// TIA Portal project "DATN" (V16) (continued)
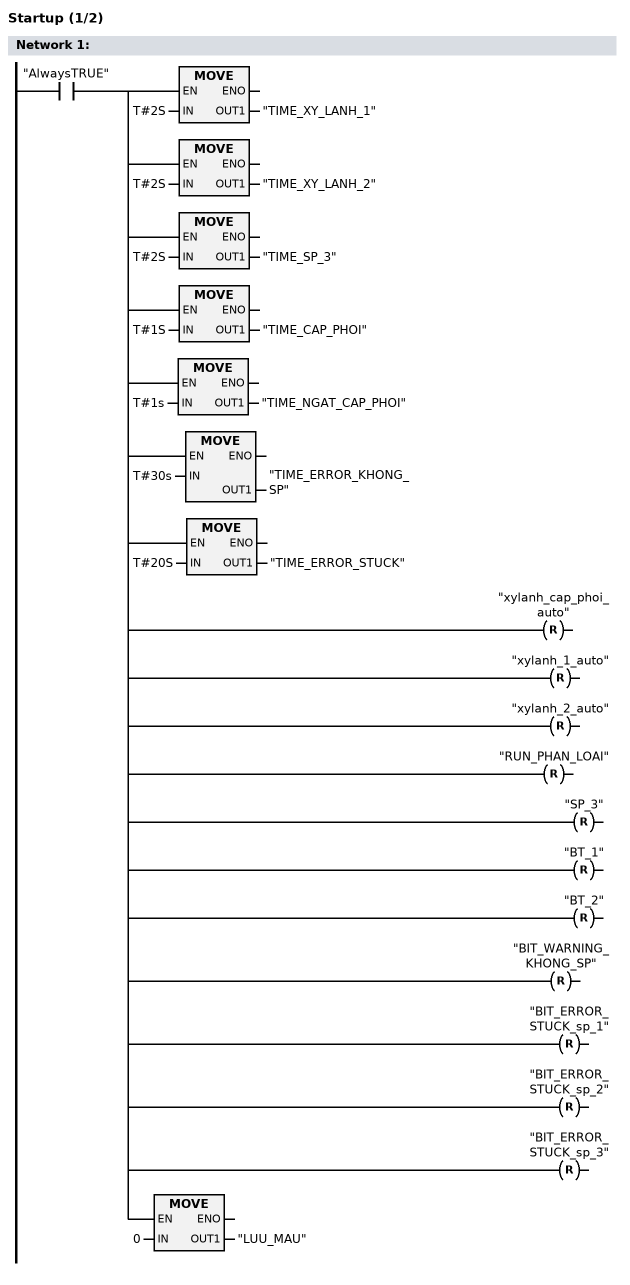
   RUNG wire#powerrail
      Contact( "AlwaysTRUE" )
      wire#w1
      Move(in := T#2S, out1 => "TIME_XY_LANH_1")
   END_RUNG
   RUNG wire#w1
      Move(in := T#2S, out1 => "TIME_XY_LANH_2")
   END_RUNG
   RUNG wire#w1
      Move(in := T#2S, out1 => "TIME_SP_3")
   END_RUNG
   RUNG wire#w1
      Move(in := T#1S, out1 => "TIME_CAP_PHOI")
   END_RUNG
   RUNG wire#w1
      Move(in := T#1s, out1 => "TIME_NGAT_CAP_PHOI")
   END_RUNG
   RUNG wire#w1
      Move(in := T#30s, out1 => "TIME_ERROR_KHONG_SP")
   END_RUNG
   RUNG wire#w1
      Move(in := T#20S, out1 => "TIME_ERROR_STUCK")
   END_RUNG
   RUNG wire#w1
      R_Coil( "xylanh_cap_phoi_auto" )
   END_RUNG
   RUNG wire#w1
      R_Coil( "xylanh_1_auto" )
   END_RUNG
   RUNG wire#w1
      R_Coil( "xylanh_2_auto" )
   END_RUNG
   RUNG wire#w1
      R_Coil( "RUN_PHAN_LOAI" )
   END_RUNG
   RUNG wire#w1
      R_Coil( "SP_3" )
   END_RUNG
   RUNG wire#w1
      R_Coil( "BT_1" )
   END_RUNG
   RUNG wire#w1
      R_Coil( "BT_2" )
   END_RUNG
   RUNG wire#w1
      R_Coil( "BIT_WARNING_KHONG_SP" )
   END_RUNG
   RUNG wire#w1
      R_Coil( "BIT_ERROR_STUCK_sp_1" )
   END_RUNG
   RUNG wire#w1
      R_Coil( "BIT_ERROR_STUCK_sp_2" )
   END_RUNG
   RUNG wire#w1
      R_Coil( "BIT_ERROR_STUCK_sp_3" )
   END_RUNG
   RUNG wire#w1
      Move(in := 0, out1 => "LUU_MAU")
   END_RUNG
   // the same network as SCL:
   IF "AlwaysTRUE" THEN
       "TIME_XY_LANH_1" := T#2S;
       "TIME_XY_LANH_2" := T#2S;
       "TIME_SP_3" := T#2S;
       "TIME_CAP_PHOI" := T#1S;
       "TIME_NGAT_CAP_PHOI" := T#1s;
       "TIME_ERROR_KHONG_SP" := T#30s;
       "TIME_ERROR_STUCK" := T#20S;
       "xylanh_cap_phoi_auto" := FALSE;
       "xylanh_1_auto" := FALSE;
       "xylanh_2_auto" := FALSE;
       "RUN_PHAN_LOAI" := FALSE;
       "SP_3" := FALSE;
       "BT_1" := FALSE;
       "BT_2" := FALSE;
       "BIT_WARNING_KHONG_SP" := FALSE;
       "BIT_ERROR_STUCK_sp_1" := FALSE;
       "BIT_ERROR_STUCK_sp_2" := FALSE;
       "BIT_ERROR_STUCK_sp_3" := FALSE;
       "LUU_MAU" := 0;
   END_IF;
END_REGION

REGION Network 2
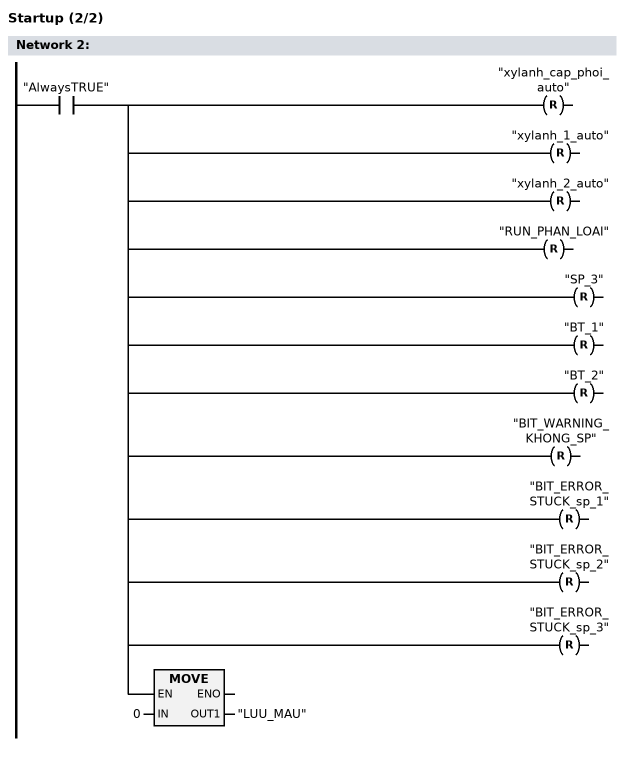
   RUNG wire#powerrail
      Contact( "AlwaysTRUE" )
      wire#w1
      R_Coil( "xylanh_cap_phoi_auto" )
   END_RUNG
   RUNG wire#w1
      R_Coil( "xylanh_1_auto" )
   END_RUNG
   RUNG wire#w1
      R_Coil( "xylanh_2_auto" )
   END_RUNG
   RUNG wire#w1
      R_Coil( "RUN_PHAN_LOAI" )
   END_RUNG
   RUNG wire#w1
      R_Coil( "SP_3" )
   END_RUNG
   RUNG wire#w1
      R_Coil( "BT_1" )
   END_RUNG
   RUNG wire#w1
      R_Coil( "BT_2" )
   END_RUNG
   RUNG wire#w1
      R_Coil( "BIT_WARNING_KHONG_SP" )
   END_RUNG
   RUNG wire#w1
      R_Coil( "BIT_ERROR_STUCK_sp_1" )
   END_RUNG
   RUNG wire#w1
      R_Coil( "BIT_ERROR_STUCK_sp_2" )
   END_RUNG
   RUNG wire#w1
      R_Coil( "BIT_ERROR_STUCK_sp_3" )
   END_RUNG
   RUNG wire#w1
      Move(in := 0, out1 => "LUU_MAU")
   END_RUNG
   // the same network as SCL:
   IF "AlwaysTRUE" THEN
       "xylanh_cap_phoi_auto" := FALSE;
       "xylanh_1_auto" := FALSE;
       "xylanh_2_auto" := FALSE;
       "RUN_PHAN_LOAI" := FALSE;
       "SP_3" := FALSE;
       "BT_1" := FALSE;
       "BT_2" := FALSE;
       "BIT_WARNING_KHONG_SP" := FALSE;
       "BIT_ERROR_STUCK_sp_1" := FALSE;
       "BIT_ERROR_STUCK_sp_2" := FALSE;
       "BIT_ERROR_STUCK_sp_3" := FALSE;
       "LUU_MAU" := 0;
   END_IF;
END_REGION
END_ORGANIZATION_BLOCK

(* ===== HMI "HMI_RT_1" =====
system functions are stored by id; their names below are inferred from use
connection "HMI_Connection_1": ETHERNET, S7_1200_OMS

HMI tags "Default tag table"
   "HMI_PB_START" : Bool = PLC HMI_PB_START AT %M100.4, 1 s
   "HMI_PB_STOP" : Bool = PLC HMI_PB_STOP AT %M100.5, 1 s
   "HMI_PB_RESET" : Bool = PLC HMI_PB_RESET AT %M100.6, 1 s
   "DEN_START" : Bool = PLC DEN_START AT %Q0.5, 1 s
   "DEN_STOP" : Bool = PLC DEN_STOP AT %Q0.6, 1 s
   "DEN_RESET" : Bool = PLC DEN_RESET AT %Q0.7, 1 s
   "HMI_AUTO_MAN" : Bool = PLC HMI_AUTO_MAN AT %M101.3, 1 s
   "COUNTER_SP_1_CV" : Int = PLC COUNTER_SP_1.CV, 1 s
   "COUNTER_SP_2_CV" : Int = PLC COUNTER_SP_2.CV, 1 s
   "COUNTER_SP_3_CV" : Int = PLC COUNTER_SP_3.CV, 1 s
   "gh_sp_GH_SP_1" : USInt = PLC gh_sp.GH_SP_1, 1 s
   "gh_sp_GH_SP_2" : USInt = PLC gh_sp.GH_SP_2, 1 s
   "gh_sp_GH_SP_3" : USInt = PLC gh_sp.GH_SP_3, 1 s
   "BANG_TAI" : Bool = PLC BANG_TAI AT %Q0.0, 1 s
   "XY_LANH_2" : Bool = PLC XY_LANH_2 AT %Q0.2, 1 s
   "XY_LANH_1" : Bool = PLC XY_LANH_1 AT %Q0.1, 1 s
   "Mau Sac" : Int = PLC "Mau Sac" AT %MW220, 1 s
   "CB_SP_2" : Bool = PLC CB_SP_2 AT %I0.2, 1 s
   "CB_SP_1" : Bool = PLC CB_SP_1 AT %I0.1, 1 s
   "CB_SP_3" : Bool = PLC CB_SP_3 AT %I0.3, 1 s
   "CB_CAP_PHOI" : Bool = PLC CB_CAP_PHOI AT %I0.0, 1 s
   "XY_LANH_CAP_PHOI_1" : Bool = PLC XY_LANH_CAP_PHOI_1 AT %Q0.3, 1 s
   "MODE_AUTO" : Bool = PLC MODE_AUTO AT %M201.7, 1 s
   "MODE_MAN" : Bool = PLC MODE_MAN AT %M202.0, 1 s
   "MAN_BT" : Bool = PLC MAN_BT AT %M100.7, 1 s
   "MAN_CAP_PHOI" : Bool = PLC MAN_CAP_PHOI AT %M101.2, 1 s
   "MAN_XYLANH_1" : Bool = PLC MAN_XYLANH_1 AT %M101.0, 1 s
   "MAN_XYLANH_2" : Bool = PLC MAN_XYLANH_2 AT %M101.1, 1 s
   "OUT_counter_1" : Bool = PLC OUT_counter_1 AT %M201.4, 1 s
   "OUT_counter_2" : Bool = PLC OUT_counter_2 AT %M201.5, 1 s
   "OUT_counter_3" : Bool = PLC OUT_counter_3 AT %M201.6, 1 s
   "RST_SP_3" : Bool = PLC RST_SP_3 AT %M101.6, 1 s
   "RST_SP_2" : Bool = PLC RST_SP_2 AT %M101.5, 1 s
   "RST_SP_1" : Bool = PLC RST_SP_1 AT %M101.4, 1 s
   "LUU_MAU" : Int = PLC LUU_MAU AT %MW222, 1 s
   "MULTI_ERROR" : Bool = PLC MULTI_ERROR AT %M450.0, 1 s
   "BIT_WARNING_KHONG_SP" : Bool = PLC BIT_WARNING_KHONG_SP AT %M400.0, 1 s
   "BIT_ERROR_STUCK_sp_1" : Bool = PLC BIT_ERROR_STUCK_sp_1 AT %M402.0, 1 s
   "BIT_ERROR_STUCK_sp_2" : Bool = PLC BIT_ERROR_STUCK_sp_2 AT %M404.0, 1 s
   "BIT_ERROR_STUCK_sp_3" : Bool = PLC BIT_ERROR_STUCK_sp_3 AT %M406.0, 1 s

HMI tags "HMI_ALARM"
   "DATA_WARNING" : Int = PLC DATA_WORD_WARNING AT %MW400, 1 s
   "DATA_ERROR_1" : Int = PLC DATA_WORD_ERROR_1 AT %MW402, 1 s
   "DATA_ERROR_2" : Int = PLC DATA_WORD_ERROR_2 AT %MW404, 1 s
   "DATA_ERROR_3" : Int = PLC DATA_WORD_ERROR_3 AT %MW406, 1 s

discrete alarms
   4: 'Cảnh báo không có sản phẩm', class Warnings, trigger "DATA_WARNING" bit 8
   1: 'Lỗi kẹt sản phẩm 1', class Warnings, trigger "DATA_ERROR_1" bit 8
   2: 'Lỗi kẹt sản phẩm 2', class Warnings, trigger "DATA_ERROR_2" bit 8
   3: 'Lỗi kẹt sản phẩm 3', class Warnings, trigger "DATA_ERROR_3" bit 8

screen "1_Login" 1440x900
   GraphicView "Graphic view_4" at 0,0 size 1438x897; Picture "plc"
   Button "Button_1" at 1010,602 size 237x78; TextOff 'LOG IN'; TextOn '2_Home'; Authorization "Operate"
      on Click: ActivateScreen("2_Home", 0)

screen "2_Home" 1440x900
   Circle "Circle_8" at 525,299 size 20x20
      Visibility <- "XY_LANH_2"
   Group "Group_7" at 531,249 size 89x62
   Polyline "Polyline_1" at 532,284 size 40x22
      Visibility <- "XY_LANH_2"
   Polyline "Polyline_2" at 531,249 size 89x62
      Visibility <- "XY_LANH_2"
   Group "Group_8" at 525,249 size 95x70
   Circle "Circle_9" at 525,299 size 20x20
      Visibility <- "XY_LANH_2"
   Circle "Circle_10" at 773,299 size 20x20
      Visibility <- "XY_LANH_1"
   Group "Group_9" at 779,249 size 89x62
   Polyline "Polyline_3" at 780,284 size 40x22
      Visibility <- "XY_LANH_1"
   Polyline "Polyline_4" at 779,249 size 89x62
      Visibility <- "XY_LANH_1"
   Group "Group_10" at 773,249 size 95x70
   Circle "Circle_11" at 773,299 size 20x20
      Visibility <- "XY_LANH_1"
   SymbolLibrary "Symbol library_14" at 1038,320 size 72x64
      Visibility <- "LUU_MAU"
   GraphicView "Graphic view_1" at 1039,340 size 58x29; Picture "Graphic_2"
      Visibility <- "LUU_MAU"
   SymbolLibrary "Symbol library_13" at 1020,330 size 72x64
      Visibility <- "LUU_MAU"
   GraphicView "Graphic view_3" at 1021,348 size 58x33; Picture "Graphic_4"
      Visibility <- "LUU_MAU"
   SymbolLibrary "Symbol library_12" at 1002,342 size 72x64
      Visibility <- "LUU_MAU"
   GraphicView "Graphic view_2" at 1003,360 size 58x33; Picture "Graphic_5"
      Visibility <- "LUU_MAU"
   SymbolLibrary "Symbol library_21" at 349,368 size 17x150
   SymbolLibrary "Symbol library_6" at 93,426 size 168x95
      Appearance <- "OUT_counter_3"
   SymbolLibrary "Symbol library_17" at 333,345 size 56x52
   SymbolLibrary "Symbol library_20" at 1179,373 size 17x150
   SymbolLibrary "Symbol library_16" at 1161,350 size 56x52
   SymbolLibrary "Symbol library_1" at 242,368 size 545x73
      Appearance <- "BANG_TAI"
   SymbolLibrary "Symbol library_2" at 650,368 size 545x73
      Appearance <- "BANG_TAI"
   SymbolLibrary "Symbol library_19" at 1082,432 size 17x150
   Group "Group_6" at 595,168 size 143x104
   Group "Group_12" at 525,249 size 95x70
   Group "Group_1" at 843,168 size 143x104
   Group "Group_11" at 773,249 size 95x70
   SymbolLibrary "Symbol library_4" at 334,546 size 168x95
      Appearance <- "OUT_counter_2"
   SymbolLibrary "Symbol library_5" at 570,546 size 168x95
      Appearance <- "OUT_counter_1"
   SymbolLibrary "Symbol library_8" at 1025,248 size 55x27
      Appearance <- "Mau Sac"
   SymbolLibrary "Symbol library_10" at 649,242 size 28x55
      Appearance <- "CB_SP_2"
   SymbolLibrary "Symbol library_11" at 902,242 size 28x55
      Appearance <- "CB_SP_1"
   TextField "Text field_6" at 679,244 size 39x25; Text 'CB2'
   TextField "Text field_7" at 931,244 size 39x25; Text 'CB1'
   TextField "Text field_9" at 569,140 size 114x56; Text 'Xy lanh loại 2'
   TextField "Text field_10" at 826,140 size 114x56; Text 'Xy lanh loại 1'
   IOField "I/O field_4" at 378,594 size 62x32; FormatPattern 99999
      ProcessValue <- "COUNTER_SP_2_CV"
   IOField "I/O field_5" at 614,594 size 62x32; FormatPattern 99999
      ProcessValue <- "COUNTER_SP_1_CV"
   TextField "Text field_14" at 103,514 size 123x43; Text 'SP Loại 3'
   TextField "Text field_15" at 456,605 size 123x43; Text 'SP Loại 2'
   TextField "Text field_16" at 693,605 size 123x43; Text 'SP Loại 1'
   Group "Group_15" at 1038,320 size 72x64; Picture "Graphic_2"
   Group "Group_16" at 1020,330 size 72x64; Picture "Graphic_4"
   SymbolLibrary "Symbol library_15" at 1065,403 size 56x52
   TextField "Text field_17" at 899,520 size 138x61; Text 'ĐỘNG CƠ BĂNG TẢI'
   Group "Group_17" at 1002,342 size 72x64; Picture "Graphic_5"
   Group "Group_13" at 385,415 size 133x122
   SymbolLibrary "Symbol library_3" at 928,463 size 110x66
      Appearance <- "BANG_TAI"
   IOField "I/O field_6" at 137,480 size 62x32; FormatPattern 99999
      ProcessValue <- "COUNTER_SP_3_CV"
   SymbolLibrary "Symbol library_22" at 243,427 size 17x150
   SymbolLibrary "Symbol library_18" at 225,404 size 56x52
   Group "Group_2" at 625,415 size 133x122
   Button "Button_3" at 11,123 size 112x37; TextOff 'Home'
      on Click: ActivateScreen("2_Home", 0)
   Button "Button_4" at 11,177 size 112x37; TextOff 'Control'; Authorization "User administration"
      on Click: ActivateScreen("3_Control", 0)
   Button "Button_6" at 11,285 size 112x37; TextOff 'Log out'
      on Click: function_f23ef4c9(); ActivateScreen("1_Login", 0)
   DateTimeField "Date/time field_3" at 1186,44 size 102x23
   DateTimeField "Date/time field_1" at 1186,18 size 254x23
   GraphicView "Graphic view_8" at 38,8 size 70x70; Picture "Hcmute"
   GraphicView "Graphic view_9" at 128,8 size 70x70; Picture "feee"
   TextField "Text field_3" at 261,15 size 906x70; Text 'HỆ THỐNG PHÂN LOẠI SẢN PHẨM THEO MÀU SẮC DÙNG XỬ LÝ ẢNH'
   GraphicView "Graphic view_10" at 134,130 size 36x18; Picture "Graphic_17"
   TextField "Text field_1" at 250,147 size 15x22; Text 'Text'
   TextField "Text field_4" at 72,730 size 139x22; Text 'Hệ thống nút nhấn'
   Button "Button_1" at 26,801 size 64x64; TextOff 'Text'; PictureOff "3-D green button (not pressed)_3"; PictureOn "3-D green button (pressed)_2"
      on Press: SetBit("HMI_PB_START")
      on Release: ResetBit("HMI_PB_START")
   TextField "Text field_5" at 31,768 size 54x22; Text 'START'
   TextField "Text field_8" at 353,730 size 133x22; Text 'Hệ thống đèn báo'
   Button "Button_2" at 109,801 size 64x64; TextOff 'Text'; PictureOff "3-D red button (not pressed)"; PictureOn "3-D red button (pressed)"
      on Press: SetBit("HMI_PB_STOP")
      on Release: ResetBit("HMI_PB_STOP")
   TextField "Text field_11" at 118,768 size 46x22; Text 'STOP'
   Button "Button_7" at 193,801 size 64x64; TextOff 'Text'; PictureOff "3-D yellow button (not pressed)"; PictureOn "3-D yellow button (pressed)"
      on Press: SetBit("HMI_PB_RESET")
      on Release: ResetBit("HMI_PB_RESET")
   TextField "Text field_12" at 199,768 size 53x22; Text 'RESET'
   GraphicView "Graphic view_4" at 387,801 size 64x64; Picture "Graphic_11"
      Visibility <- "DEN_STOP"
   GraphicView "Graphic view_5" at 304,801 size 64x64; Picture "Graphic_9"
      Visibility <- "DEN_START"
   GraphicView "Graphic view_6" at 471,801 size 64x64; Picture "Graphic_18"
      Visibility <- "DEN_RESET"
   GraphicView "Graphic view_7" at 304,801 size 64x64; Picture "Graphic_10"
      Visibility <- "DEN_START"
   GraphicView "Graphic view_11" at 387,801 size 64x64; Picture "Graphic_12"
      Visibility <- "DEN_STOP"
   GraphicView "Graphic view_12" at 471,801 size 64x64; Picture "Graphic_19"
      Visibility <- "DEN_RESET"
   TextField "Text field_13" at 322,768 size 29x22; Text 'ON'
   TextField "Text field_18" at 402,768 size 35x22; Text 'OFF'
   TextField "Text field_19" at 456,768 size 95x22; Text 'WARNNING'
   TextField "Text field_20" at 659,683 size 123x22; Text 'Bảng điều khiển'
   TextField "Text field_2" at 581,730 size 132x22; Text 'Chế độ hoạt động'
   Switch "Switch_1" at 587,805 size 120x60; CaptionText 'Switch'; TextOff 'OFF'; TextOn 'ON'; PictureOn "Illuminated red-green (Red)_1"; PictureOff "Illuminated red-green (Green)_1"
      ProcessValue <- "HMI_AUTO_MAN"
   TextField "Text field_23" at 973,730 size 148x22; Text 'Thông tin sản phẩm'
   TextField "Text field_24" at 895,754 size 137x22; Text 'Giới hạn số lượng'
   TextField "Text field_25" at 760,784 size 123x22; Text 'Sản phẩm loại 1'
   TextField "Text field_26" at 760,816 size 123x22; Text 'Sản phẩm loại 2'
   TextField "Text field_27" at 760,848 size 123x22; Text 'Sản phẩm loại 3'
   IOField "I/O field_1" at 916,779 size 96x32; FormatPattern 999
      ProcessValue <- "gh_sp_GH_SP_1"
   IOField "I/O field_2" at 916,811 size 96x32; FormatPattern 999
      ProcessValue <- "gh_sp_GH_SP_2"
   IOField "I/O field_3" at 916,843 size 96x32; FormatPattern 999
      ProcessValue <- "gh_sp_GH_SP_3"
   TextField "Text field_28" at 1084,754 size 130x22; Text 'Số lượng hiện tại'
   IOField "I/O field_7" at 1101,779 size 96x32; FormatPattern 99999
      ProcessValue <- "COUNTER_SP_1_CV"
   IOField "I/O field_8" at 1101,811 size 96x32; FormatPattern 99999
      ProcessValue <- "COUNTER_SP_2_CV"
   IOField "I/O field_9" at 1101,843 size 96x32; FormatPattern 99999
      ProcessValue <- "COUNTER_SP_3_CV"
   GraphicView "Graphic view_13" at 1023,406 size 94x98; Picture "Graphic_20"
   SymbolLibrary "Symbol library_7" at 349,242 size 28x55
      Appearance <- "CB_SP_3"
   TextField "Text field_29" at 385,244 size 39x25; Text 'CB3'
   SymbolLibrary "Symbol library_23" at 1215,367 size 17x155
   SymbolLibrary "Symbol library_24" at 1118,426 size 17x156
   SymbolLibrary "Symbol library_25" at 1302,367 size 17x154
   SymbolLibrary "Symbol library_26" at 1205,426 size 17x155
   SymbolLibrary "Symbol library_27" at 1183,330 size 72x64
      Visibility <- "CB_CAP_PHOI"
   SymbolLibrary "Symbol library_28" at 1287,316 size 55x28
      Appearance <- "CB_CAP_PHOI"
   SymbolLibrary "Symbol library_9" at 1243,351 size 130x26
      Visibility <- "XY_LANH_CAP_PHOI_1"
   SymbolLibrary "Symbol library_29" at 1292,351 size 82x26
      Visibility <- "XY_LANH_CAP_PHOI_1"
   TextField "Text field_30" at 1270,281 size 117x25; Text 'CB CẤP PHÔI'
   TextField "Text field_31" at 1258,754 size 134x22; Text 'Reset thùng hàng'
   Button "Button_8" at 1277,779 size 96x32; TextOff 'RST_1'
      Appearance <- "OUT_counter_1"
      on Press: SetBit("RST_SP_1")
      on Release: ResetBit("RST_SP_1")
   Button "Button_9" at 1277,810 size 96x32; TextOff 'RST_2'
      Appearance <- "OUT_counter_2"
      on Press: SetBit("RST_SP_2")
      on Release: ResetBit("RST_SP_2")
   Button "Button_10" at 1277,841 size 96x32; TextOff 'RST_3'
      Appearance <- "OUT_counter_3"
      on Press: SetBit("RST_SP_3")
      on Release: ResetBit("RST_SP_3")
   Button "Button_5" at 11,231 size 112x37; TextOff 'Alarm'
      on Click: ActivateScreen("4_ALARM", 0)
      Appearance <- "MULTI_ERROR"
   Rectangle "Rectangle_9" at 579,754 size 65x48
      Appearance <- "MODE_AUTO"
   Rectangle "Rectangle_10" at 650,754 size 65x48
      Appearance <- "MODE_MAN"
   TextField "Text field_32" at 1203,96 size 125x22; Text 'Màu sắc hiện tại'
   Rectangle "Rectangle_13" at 1246,137 size 40x37
      Appearance <- "LUU_MAU"
   TextField "Text field_33" at 1245,185 size 42x22; Text 'Vàng'
      Visibility <- "LUU_MAU"
   TextField "Text field_34" at 1248,185 size 36x22; Text 'Lam'
      Visibility <- "LUU_MAU"
   TextField "Text field_35" at 1250,185 size 32x22; Text 'Tím'
      Visibility <- "LUU_MAU"
   TextField "Text field_36" at 1231,185 size 70x22; Text 'No Color'
      Visibility <- "LUU_MAU"
   TextField "Text field_21" at 592,768 size 39x22; Text 'Auto'
   TextField "Text field_22" at 653,768 size 59x22; Text 'Manual'

screen "3_Control" 1440x900
   Circle "Circle_8" at 525,299 size 20x20
      Visibility <- "XY_LANH_2"
   Group "Group_7" at 531,249 size 89x62
   Polyline "Polyline_1" at 532,284 size 40x22
      Visibility <- "XY_LANH_2"
   Polyline "Polyline_2" at 531,249 size 89x62
      Visibility <- "XY_LANH_2"
   Group "Group_8" at 525,249 size 95x70
   Circle "Circle_9" at 525,299 size 20x20
      Visibility <- "XY_LANH_2"
   Circle "Circle_10" at 773,299 size 20x20
      Visibility <- "XY_LANH_1"
   Group "Group_9" at 779,249 size 89x62
   Polyline "Polyline_3" at 780,284 size 40x22
      Visibility <- "XY_LANH_1"
   Polyline "Polyline_4" at 779,249 size 89x62
      Visibility <- "XY_LANH_1"
   Group "Group_10" at 773,249 size 95x70
   Circle "Circle_11" at 773,299 size 20x20
      Visibility <- "XY_LANH_1"
   SymbolLibrary "Symbol library_6" at 93,426 size 168x95
      Appearance <- "OUT_counter_3"
   SymbolLibrary "Symbol library_4" at 334,546 size 168x95
      Appearance <- "OUT_counter_2"
   SymbolLibrary "Symbol library_5" at 570,546 size 168x95
      Appearance <- "OUT_counter_1"
   SymbolLibrary "Symbol library_21" at 349,368 size 17x150
   SymbolLibrary "Symbol library_17" at 333,345 size 56x52
   SymbolLibrary "Symbol library_20" at 1179,373 size 17x150
   SymbolLibrary "Symbol library_16" at 1161,350 size 56x52
   SymbolLibrary "Symbol library_1" at 242,368 size 545x73
      Appearance <- "BANG_TAI"
   SymbolLibrary "Symbol library_2" at 650,368 size 545x73
      Appearance <- "BANG_TAI"
   SymbolLibrary "Symbol library_19" at 1082,432 size 17x150
   Group "Group_6" at 595,168 size 143x104
   Group "Group_12" at 525,249 size 95x70
   Group "Group_1" at 843,168 size 143x104
   Group "Group_11" at 773,249 size 95x70
   SymbolLibrary "Symbol library_8" at 1025,248 size 55x27
      Appearance <- "Mau Sac"
   SymbolLibrary "Symbol library_10" at 649,242 size 28x55
      Appearance <- "CB_SP_2"
   SymbolLibrary "Symbol library_11" at 902,242 size 28x55
      Appearance <- "CB_SP_1"
   TextField "Text field_6" at 679,244 size 39x25; Text 'CB2'
   TextField "Text field_7" at 931,244 size 39x25; Text 'CB1'
   TextField "Text field_9" at 569,140 size 114x56; Text 'Xy lanh loại 2'
   TextField "Text field_10" at 826,140 size 114x56; Text 'Xy lanh loại 1'
   IOField "I/O field_4" at 378,594 size 62x32; FormatPattern 99999
      ProcessValue <- "COUNTER_SP_2_CV"
   IOField "I/O field_5" at 614,594 size 62x32; FormatPattern 99999
      ProcessValue <- "COUNTER_SP_1_CV"
   TextField "Text field_14" at 103,514 size 123x43; Text 'SP Loại 3'
   TextField "Text field_15" at 456,605 size 123x43; Text 'SP Loại 2'
   TextField "Text field_16" at 693,605 size 123x43; Text 'SP Loại 1'
   SymbolLibrary "Symbol library_15" at 1065,403 size 56x52
   TextField "Text field_17" at 899,520 size 138x61; Text 'ĐỘNG CƠ BĂNG TẢI'
   Group "Group_13" at 385,415 size 133x122
   SymbolLibrary "Symbol library_3" at 928,463 size 110x66
      Appearance <- "BANG_TAI"
   IOField "I/O field_6" at 137,480 size 62x32; FormatPattern 99999
      ProcessValue <- "COUNTER_SP_3_CV"
   SymbolLibrary "Symbol library_22" at 243,427 size 17x150
   SymbolLibrary "Symbol library_18" at 225,404 size 56x52
   Group "Group_2" at 625,415 size 133x122
   Button "Button_3" at 11,123 size 112x37; TextOff 'Home'
      on Click: ActivateScreen("2_Home", 0)
   Button "Button_4" at 11,177 size 112x37; TextOff 'Control'
      on Click: ActivateScreen("3_Control", 0)
   Button "Button_6" at 11,285 size 112x37; TextOff 'Log out'
      on Click: ActivateScreen("1_Login", 0)
   DateTimeField "Date/time field_3" at 1186,44 size 102x23
   DateTimeField "Date/time field_1" at 1186,18 size 254x23
   GraphicView "Graphic view_8" at 38,8 size 70x70; Picture "Hcmute"
   GraphicView "Graphic view_9" at 128,8 size 70x70; Picture "feee"
   GraphicView "Graphic view_10" at 134,187 size 36x18; Picture "Graphic_17"
   TextField "Text field_1" at 250,147 size 15x22; Text 'Text'
   TextField "Text field_4" at 72,730 size 139x22; Text 'Hệ thống nút nhấn'
   Button "Button_1" at 26,801 size 64x64; TextOff 'Text'; PictureOn "3-D green button (pressed)_2"; PictureOff "3-D green button (not pressed)_3"
      on Release: ResetBit("HMI_PB_START")
      on Press: SetBit("HMI_PB_START")
   TextField "Text field_5" at 31,768 size 54x22; Text 'START'
   TextField "Text field_8" at 353,730 size 133x22; Text 'Hệ thống đèn báo'
   Button "Button_2" at 109,801 size 64x64; TextOff 'Text'; PictureOn "3-D red button (pressed)"; PictureOff "3-D red button (not pressed)"
      on Release: ResetBit("HMI_PB_STOP")
      on Press: SetBit("HMI_PB_STOP")
   TextField "Text field_11" at 118,768 size 46x22; Text 'STOP'
   Button "Button_7" at 193,801 size 64x64; TextOff 'Text'; PictureOn "3-D yellow button (pressed)"; PictureOff "3-D yellow button (not pressed)"
      on Release: ResetBit("HMI_PB_RESET")
      on Press: SetBit("HMI_PB_RESET")
   TextField "Text field_12" at 199,768 size 53x22; Text 'RESET'
   GraphicView "Graphic view_4" at 387,801 size 64x64; Picture "Graphic_11"
      Visibility <- "DEN_STOP"
   GraphicView "Graphic view_5" at 304,801 size 64x64; Picture "Graphic_9"
      Visibility <- "DEN_START"
   GraphicView "Graphic view_6" at 471,801 size 64x64; Picture "Graphic_18"
      Visibility <- "DEN_RESET"
   GraphicView "Graphic view_7" at 304,801 size 64x64; Picture "Graphic_10"
      Visibility <- "DEN_START"
   GraphicView "Graphic view_11" at 387,801 size 64x64; Picture "Graphic_12"
      Visibility <- "DEN_STOP"
   GraphicView "Graphic view_12" at 471,801 size 64x64; Picture "Graphic_19"
      Visibility <- "DEN_RESET"
   TextField "Text field_13" at 322,768 size 29x22; Text 'ON'
   TextField "Text field_18" at 402,768 size 35x22; Text 'OFF'
   TextField "Text field_19" at 456,768 size 95x22; Text 'WARNNING'
   TextField "Text field_20" at 659,683 size 123x22; Text 'Bảng điều khiển'
   TextField "Text field_2" at 581,730 size 132x22; Text 'Chế độ hoạt động'
   Switch "Switch_1" at 587,805 size 120x60; CaptionText 'Switch'; TextOff 'OFF'; TextOn 'ON'; PictureOff "Illuminated red-green (Green)_1"; PictureOn "Illuminated red-green (Red)_1"
      ProcessValue <- "HMI_AUTO_MAN"
   TextField "Text field_23" at 746,730 size 261x22; Text 'Cài đặt giới hạn số lượng sản phẩm'
   TextField "Text field_25" at 745,784 size 123x22; Text 'Sản phẩm loại 1'
   TextField "Text field_26" at 745,816 size 123x22; Text 'Sản phẩm loại 2'
   TextField "Text field_27" at 745,848 size 123x22; Text 'Sản phẩm loại 3'
   IOField "I/O field_1" at 901,779 size 96x32; FormatPattern 999
      ProcessValue <- "gh_sp_GH_SP_1"
   IOField "I/O field_2" at 901,811 size 96x32; FormatPattern 999
      ProcessValue <- "gh_sp_GH_SP_2"
   IOField "I/O field_3" at 901,843 size 96x32; FormatPattern 999
      ProcessValue <- "gh_sp_GH_SP_3"
   GraphicView "Graphic view_13" at 1023,406 size 94x98; Picture "Graphic_20"
   SymbolLibrary "Symbol library_7" at 349,242 size 28x55
      Appearance <- "CB_SP_3"
   TextField "Text field_29" at 385,244 size 39x25; Text 'CB3'
   SymbolLibrary "Symbol library_23" at 1215,367 size 17x155
   SymbolLibrary "Symbol library_24" at 1118,426 size 17x156
   SymbolLibrary "Symbol library_25" at 1302,367 size 17x154
   SymbolLibrary "Symbol library_26" at 1205,426 size 17x155
   SymbolLibrary "Symbol library_27" at 1183,330 size 72x64
      Visibility <- "CB_CAP_PHOI"
   SymbolLibrary "Symbol library_28" at 1287,316 size 55x28
      Appearance <- "CB_CAP_PHOI"
   SymbolLibrary "Symbol library_9" at 1243,351 size 130x26
      Visibility <- "XY_LANH_CAP_PHOI_1"
   SymbolLibrary "Symbol library_29" at 1292,351 size 82x26
      Visibility <- "XY_LANH_CAP_PHOI_1"
   TextField "Text field_30" at 1270,281 size 117x25; Text 'CB CẤP PHÔI'
   Rectangle "Rectangle_9" at 579,754 size 65x48
      Appearance <- "MODE_AUTO"
   Rectangle "Rectangle_10" at 650,754 size 65x48
      Appearance <- "MODE_MAN"
   TextField "Text field_21" at 592,768 size 39x22; Text 'Auto'
   TextField "Text field_22" at 653,768 size 59x22; Text 'Manual'
   TextField "Text field_24" at 1158,730 size 153x22; Text 'Điều khiển bằng tay'
   Button "Button_8" at 1062,779 size 160x32; TextOff 'Băng tải'
      Appearance <- "BANG_TAI"
      on Press: SetBit("MAN_BT")
      on Release: ResetBit("MAN_BT")
   Button "Button_9" at 1062,843 size 160x32; TextOff 'Xylanh cấp phôi'
      Appearance <- "XY_LANH_CAP_PHOI_1"
      on Press: SetBit("MAN_CAP_PHOI")
      on Release: ResetBit("MAN_CAP_PHOI")
   Button "Button_10" at 1256,779 size 160x32; TextOff 'Xylanh 1'
      Appearance <- "XY_LANH_1"
      on Press: SetBit("MAN_XYLANH_1")
      on Release: ResetBit("MAN_XYLANH_1")
   Button "Button_11" at 1256,843 size 160x32; TextOff 'Xylanh 2'
      Appearance <- "XY_LANH_2"
      on Press: SetBit("MAN_XYLANH_2")
      on Release: ResetBit("MAN_XYLANH_2")
   Button "Button_5" at 11,231 size 112x37; TextOff 'Alarm'
      on Click: ActivateScreen("4_ALARM", 0)
      Appearance <- "MULTI_ERROR"
   TextField "Text field_32" at 1203,96 size 125x22; Text 'Màu sắc hiện tại'
   Rectangle "Rectangle_13" at 1246,137 size 40x37
      Appearance <- "LUU_MAU"
   TextField "Text field_33" at 1245,185 size 42x22; Text 'Vàng'
      Visibility <- "LUU_MAU"
   TextField "Text field_34" at 1248,185 size 36x22; Text 'Lam'
      Visibility <- "LUU_MAU"
   TextField "Text field_35" at 1250,185 size 32x22; Text 'Tím'
      Visibility <- "LUU_MAU"
   TextField "Text field_36" at 1231,185 size 70x22; Text 'No Color'
      Visibility <- "LUU_MAU"
   Group "Group_15" at 1038,320 size 72x64; Picture "Graphic_2"
   Group "Group_16" at 1020,330 size 72x64; Picture "Graphic_4"
   Group "Group_17" at 1002,342 size 72x64; Picture "Graphic_5"
   TextField "Text field_3" at 261,15 size 906x70; Text 'HỆ THỐNG PHÂN LOẠI SẢN PHẨM THEO MÀU SẮC DÙNG XỬ LÝ ẢNH'
   SymbolLibrary "Symbol library_14" at 1038,320 size 72x64
      Visibility <- "LUU_MAU"
   GraphicView "Graphic view_1" at 1039,340 size 58x29; Picture "Graphic_2"
      Visibility <- "LUU_MAU"
   SymbolLibrary "Symbol library_13" at 1020,330 size 72x64
      Visibility <- "LUU_MAU"
   GraphicView "Graphic view_3" at 1021,348 size 58x33; Picture "Graphic_4"
      Visibility <- "LUU_MAU"
   SymbolLibrary "Symbol library_12" at 1002,342 size 72x64
      Visibility <- "LUU_MAU"
   GraphicView "Graphic view_2" at 1003,360 size 58x33; Picture "Graphic_5"
      Visibility <- "LUU_MAU"

screen "4_ALARM" 1440x900
   SymbolLibrary "Symbol library_21" at 349,368 size 17x150
   SymbolLibrary "Symbol library_6" at 93,426 size 168x95
      Appearance <- "OUT_counter_3"
   SymbolLibrary "Symbol library_17" at 333,345 size 56x52
   SymbolLibrary "Symbol library_20" at 1179,373 size 17x150
   SymbolLibrary "Symbol library_16" at 1161,350 size 56x52
   SymbolLibrary "Symbol library_1" at 242,368 size 545x73
      Appearance <- "BANG_TAI"
   SymbolLibrary "Symbol library_2" at 650,368 size 545x73
      Appearance <- "BANG_TAI"
   SymbolLibrary "Symbol library_19" at 1082,432 size 17x150
   Group "Group_6" at 595,168 size 143x104
   Group "Group_12" at 525,249 size 95x70
   Group "Group_1" at 843,168 size 143x104
   Group "Group_11" at 773,249 size 95x70
   SymbolLibrary "Symbol library_4" at 334,546 size 168x95
      Appearance <- "OUT_counter_2"
   SymbolLibrary "Symbol library_5" at 570,546 size 168x95
      Appearance <- "OUT_counter_1"
   SymbolLibrary "Symbol library_8" at 1025,248 size 55x27
      Appearance <- "Mau Sac"
   SymbolLibrary "Symbol library_10" at 649,242 size 28x55
      Appearance <- "CB_SP_2"
   SymbolLibrary "Symbol library_11" at 902,242 size 28x55
      Appearance <- "CB_SP_1"
   TextField "Text field_6" at 679,244 size 39x25; Text 'CB2'
   TextField "Text field_7" at 931,244 size 39x25; Text 'CB1'
   TextField "Text field_9" at 569,140 size 114x56; Text 'Xy lanh loại 2'
   TextField "Text field_10" at 826,140 size 114x56; Text 'Xy lanh loại 1'
   IOField "I/O field_4" at 378,594 size 62x32; FormatPattern 99999
      ProcessValue <- "COUNTER_SP_2_CV"
   IOField "I/O field_5" at 614,594 size 62x32; FormatPattern 99999
      ProcessValue <- "COUNTER_SP_1_CV"
   TextField "Text field_14" at 103,514 size 123x43; Text 'SP Loại 3'
   TextField "Text field_15" at 456,605 size 123x43; Text 'SP Loại 2'
   TextField "Text field_16" at 693,605 size 123x43; Text 'SP Loại 1'
   SymbolLibrary "Symbol library_15" at 1065,403 size 56x52
   TextField "Text field_17" at 899,520 size 138x61; Text 'ĐỘNG CƠ BĂNG TẢI'
   Group "Group_13" at 385,415 size 133x122
   SymbolLibrary "Symbol library_3" at 928,463 size 110x66
      Appearance <- "BANG_TAI"
   IOField "I/O field_6" at 137,480 size 62x32; FormatPattern 99999
      ProcessValue <- "COUNTER_SP_3_CV"
   SymbolLibrary "Symbol library_22" at 243,427 size 17x150
   SymbolLibrary "Symbol library_18" at 225,404 size 56x52
   Group "Group_2" at 625,415 size 133x122
   Button "Button_3" at 11,123 size 112x37; TextOff 'Home'
      on Click: ActivateScreen("2_Home", 0)
   Button "Button_4" at 11,177 size 112x37; TextOff 'Control'
      on Click: ActivateScreen("3_Control", 0)
   Button "Button_5" at 11,231 size 112x37; TextOff 'Alarm'
      on Click: ActivateScreen("4_ALARM", 0)
      Appearance <- "MULTI_ERROR"
   Button "Button_6" at 11,285 size 112x37; TextOff 'Log out'
      on Click: function_f23ef4c9(); ActivateScreen("1_Login", 0)
   DateTimeField "Date/time field_3" at 1186,44 size 102x23
   DateTimeField "Date/time field_1" at 1186,18 size 254x23
   GraphicView "Graphic view_8" at 38,8 size 70x70; Picture "Hcmute"
   GraphicView "Graphic view_9" at 128,8 size 70x70; Picture "feee"
   GraphicView "Graphic view_10" at 134,241 size 36x18; Picture "Graphic_17"
   TextField "Text field_1" at 250,147 size 15x22; Text 'Text'
   TextField "Text field_4" at 72,730 size 139x22; Text 'Hệ thống nút nhấn'
   Button "Button_1" at 26,801 size 64x64; TextOff 'Text'; PictureOn "3-D green button (pressed)_2"; PictureOff "3-D green button (not pressed)_3"
      on Release: ResetBit("HMI_PB_START")
      on Press: SetBit("HMI_PB_START")
   TextField "Text field_5" at 31,768 size 54x22; Text 'START'
   TextField "Text field_8" at 353,730 size 133x22; Text 'Hệ thống đèn báo'
   Button "Button_2" at 109,801 size 64x64; TextOff 'Text'; PictureOn "3-D red button (pressed)"; PictureOff "3-D red button (not pressed)"
      on Release: ResetBit("HMI_PB_STOP")
      on Press: SetBit("HMI_PB_STOP")
   TextField "Text field_11" at 118,768 size 46x22; Text 'STOP'
   Button "Button_7" at 193,801 size 64x64; TextOff 'Text'; PictureOn "3-D yellow button (pressed)"; PictureOff "3-D yellow button (not pressed)"
      on Release: ResetBit("HMI_PB_RESET")
      on Press: SetBit("HMI_PB_RESET")
   TextField "Text field_12" at 199,768 size 53x22; Text 'RESET'
   GraphicView "Graphic view_4" at 387,801 size 64x64; Picture "Graphic_11"
      Visibility <- "DEN_STOP"
   GraphicView "Graphic view_5" at 304,801 size 64x64; Picture "Graphic_9"
      Visibility <- "DEN_START"
   GraphicView "Graphic view_6" at 471,801 size 64x64; Picture "Graphic_18"
      Visibility <- "DEN_RESET"
   GraphicView "Graphic view_7" at 304,801 size 64x64; Picture "Graphic_10"
      Visibility <- "DEN_START"
   GraphicView "Graphic view_11" at 387,801 size 64x64; Picture "Graphic_12"
      Visibility <- "DEN_STOP"
   GraphicView "Graphic view_12" at 471,801 size 64x64; Picture "Graphic_19"
      Visibility <- "DEN_RESET"
   TextField "Text field_13" at 322,768 size 29x22; Text 'ON'
   TextField "Text field_18" at 402,768 size 35x22; Text 'OFF'
   TextField "Text field_19" at 456,768 size 95x22; Text 'WARNNING'
   TextField "Text field_20" at 659,683 size 123x22; Text 'Bảng điều khiển'
   TextField "Text field_2" at 581,730 size 132x22; Text 'Chế độ hoạt động'
   Switch "Switch_1" at 587,805 size 120x60; CaptionText 'Switch'; TextOff 'OFF'; TextOn 'ON'; PictureOff "Illuminated red-green (Green)_1"; PictureOn "Illuminated red-green (Red)_1"
      ProcessValue <- "HMI_AUTO_MAN"
   GraphicView "Graphic view_13" at 1023,406 size 94x98; Picture "Graphic_20"
   SymbolLibrary "Symbol library_7" at 349,242 size 28x55
      Appearance <- "CB_SP_3"
   TextField "Text field_29" at 385,244 size 39x25; Text 'CB3'
   SymbolLibrary "Symbol library_23" at 1215,367 size 17x155
   SymbolLibrary "Symbol library_24" at 1118,426 size 17x156
   SymbolLibrary "Symbol library_25" at 1302,367 size 17x154
   SymbolLibrary "Symbol library_26" at 1205,426 size 17x155
   Polygon "Polygon_5" at 1118,366 size 202x60
      Appearance <- "BIT_WARNING_KHONG_SP"
   SymbolLibrary "Symbol library_27" at 1183,330 size 72x64
      Visibility <- "CB_CAP_PHOI"
   SymbolLibrary "Symbol library_28" at 1287,316 size 55x28
      Appearance <- "CB_CAP_PHOI"
   SymbolLibrary "Symbol library_9" at 1243,351 size 130x26
      Visibility <- "XY_LANH_CAP_PHOI_1"
   SymbolLibrary "Symbol library_29" at 1292,351 size 82x26
      Visibility <- "XY_LANH_CAP_PHOI_1"
   TextField "Text field_30" at 1270,281 size 117x25; Text 'CB CẤP PHÔI'
   AlarmView "Alarm view_1" at 739,716 size 680x169
   Rectangle "Rectangle_9" at 579,754 size 65x48
      Appearance <- "MODE_AUTO"
   Rectangle "Rectangle_10" at 650,754 size 65x48
      Appearance <- "MODE_MAN"
   TextField "Text field_21" at 592,768 size 39x22; Text 'Auto'
   TextField "Text field_22" at 653,768 size 59x22; Text 'Manual'
   Group "Group_3" at 882,342 size 72x64; Picture "Graphic_5"
   TextField "Text field_32" at 1203,96 size 125x22; Text 'Màu sắc hiện tại'
   Rectangle "Rectangle_13" at 1246,137 size 40x37
      Appearance <- "LUU_MAU"
   TextField "Text field_33" at 1245,185 size 42x22; Text 'Vàng'
      Visibility <- "LUU_MAU"
   TextField "Text field_34" at 1248,185 size 36x22; Text 'Lam'
      Visibility <- "LUU_MAU"
   TextField "Text field_35" at 1250,185 size 32x22; Text 'Tím'
      Visibility <- "LUU_MAU"
   TextField "Text field_36" at 1231,185 size 70x22; Text 'No Color'
      Visibility <- "LUU_MAU"
   Group "Group_4" at 343,330 size 72x64; Picture "Graphic_4"
   Group "Group_5" at 643,320 size 72x64; Picture "Graphic_2"
   TextField "Text field_3" at 261,15 size 906x70; Text 'HỆ THỐNG PHÂN LOẠI SẢN PHẨM THEO MÀU SẮC DÙNG XỬ LÝ ẢNH'
   Circle "Circle_8" at 525,299 size 20x20
      Visibility <- "XY_LANH_2"
   Group "Group_7" at 531,249 size 89x62
   Polyline "Polyline_1" at 532,284 size 40x22
      Visibility <- "XY_LANH_2"
   Polyline "Polyline_2" at 531,249 size 89x62
      Visibility <- "XY_LANH_2"
   Group "Group_8" at 525,249 size 95x70
   Circle "Circle_9" at 525,299 size 20x20
      Visibility <- "XY_LANH_2"
   Circle "Circle_10" at 773,299 size 20x20
      Visibility <- "XY_LANH_1"
   Group "Group_9" at 779,249 size 89x62
   Polyline "Polyline_3" at 780,284 size 40x22
      Visibility <- "XY_LANH_1"
   Polyline "Polyline_4" at 779,249 size 89x62
      Visibility <- "XY_LANH_1"
   Group "Group_10" at 773,249 size 95x70
   Circle "Circle_11" at 773,299 size 20x20
      Visibility <- "XY_LANH_1"
   SymbolLibrary "Symbol library_30" at 882,342 size 72x64
      Visibility <- "BIT_ERROR_STUCK_sp_1"
      Appearance <- "BIT_ERROR_STUCK_sp_1"
   GraphicView "Graphic view_14" at 883,360 size 58x33; Picture "Graphic_5"
      Visibility <- "BIT_ERROR_STUCK_sp_1"
   SymbolLibrary "Symbol library_31" at 343,330 size 72x64
      Visibility <- "BIT_ERROR_STUCK_sp_3"
      Appearance <- "BIT_ERROR_STUCK_sp_3"
   GraphicView "Graphic view_15" at 344,348 size 58x33; Picture "Graphic_4"
      Visibility <- "BIT_ERROR_STUCK_sp_3"
   SymbolLibrary "Symbol library_32" at 643,320 size 72x64
      Visibility <- "BIT_ERROR_STUCK_sp_2"
      Appearance <- "BIT_ERROR_STUCK_sp_2"
   GraphicView "Graphic view_16" at 644,340 size 58x29; Picture "Graphic_2"
      Visibility <- "BIT_ERROR_STUCK_sp_2"
*)